FUNCTION_BLOCK "CPG_RecipeSetpoint_STRING"   // FB31617, SCL
TITLE = CPG_RecipeSetpoint_STRING
{ S7_Optimized_Access := 'TRUE' }
AUTHOR : tech.team.motioncontrol@siemens.com
FAMILY : CPG
VERSION : 1.1
// Support: tech.team.motioncontrol@siemens.com
   VAR_INPUT
      enable : Bool;   // If true, setpoint changes are permitted
      disableRecipeControl : Bool;   // If true, the setpoint is no longer handled as a recipe
   END_VAR
   VAR_OUTPUT
      out : String[60];   // Currently running recipe value
      changeEnabled : Bool;   // Enable input is true, setpoint can be changed
      recipeControlDisabled : Bool;   // The value is not subject to recipe controls
      changeNotAllowed : Bool;   // Change is not permitted due to machine state
      recipeSetpointDifference : Bool;   // The currently running (out) value and setpoint value are not equal
   END_VAR
   VAR_IN_OUT
      recipeControl : "CPG_typeRecipeControl";   // Recipe control tag
      recipeSetpoint : "CPG_typeRecipeSetpoint_STRING";   // Recipe setpoint tag
   END_VAR
   VAR
      statFirstScan : Bool := true;
      statPrevChangeNum : Int;
      statPrevSaveNum : Int;
      statPrevCopyNum : Int;
      statPrevDeleteNum : Int;
      statPrevOut : String[60];
      statChangeNotAllowedTimer : TON_TIME;
      statTimerEN : Bool;
   END_VAR
   VAR CONSTANT
      DELAY_TIME : Time := T#3s;
   END_VAR
BEGIN
   //============================================================================================================
   // SIEMENS AG
   // (c)Copyright 2019 All Rights Reserved
   //------------------------------------------------------------------------------------------------------------
   // Library: LCPG
   // Tested with: S7-1500 with FW version V2.1
   // Engineering: TIA Portal V14
   // Restrictions: ---
   // Requirements: S7-1500
   // Functionality: instantiate this once in the program for each recipe setpoint of STRING
   // Support: tech.team.motioncontrol@siemens.com
   //------------------------------------------------------------------------------------------------------------
   // Change log table:
   // Version       Date               Expert in charge    Changes applied
   //  01.01.00     02.01.2019         KB                  Initial Release
   //============================================================================================================
   // Function : CPG_RecipeSetpoint_STRING
   //============================================================================================================

   // Language Selection
   #recipeSetpoint.CurrentSetpointName := #recipeSetpoint.SetpointName[#recipeControl.LanguageSelection];

   //Recipe Disable Control
   #recipeSetpoint.DisableRecipeControl := #disableRecipeControl;

   //Pass through enable bit
   #recipeSetpoint.SetpointChangeEnabled := #enable;

   //Set out value to match initial one on first scan
   IF #statFirstScan THEN
       #recipeSetpoint.CurrentRecipeValue := #recipeSetpoint.RecipeValues[#recipeControl.CurrentRecipeID];
       #recipeSetpoint.OUT := #recipeSetpoint.RecipeValues[#recipeControl.CurrentRecipeID];
       #statFirstScan := false;
   END_IF;


   REGION RECIPE CONTROL
       // Recipe Control - Change, Save, Copy, Delete, Revert setpoint, Save setpoint
       IF NOT (#recipeSetpoint.DisableRecipeControl) THEN
           //Recipe Change command
           IF #recipeControl.RecipeChangeNum <> #statPrevChangeNum THEN
               #recipeSetpoint.OUT := #recipeSetpoint.RecipeValues[#recipeControl.CurrentRecipeID];
               #statPrevChangeNum := #recipeControl.RecipeChangeNum;
               // Prevents multiple commands from being executed if this instruction is not being scanned
               #statPrevSaveNum := #recipeControl.RecipeSaveNum;
               #statPrevCopyNum := #recipeControl.RecipeCopyNum;
               #statPrevDeleteNum := #recipeControl.RecipeDeleteNum;
           END_IF;
           //Recipe Save command
           IF #recipeControl.RecipeSaveNum <> #statPrevSaveNum THEN
               #recipeSetpoint.RecipeValues[#recipeControl.RecipeDestinationID] := #recipeSetpoint.OUT;
               #statPrevSaveNum := #recipeControl.RecipeSaveNum;
               // Prevents multiple commands from being executed if this instruction is not being scanned
               #statPrevCopyNum := #recipeControl.RecipeCopyNum;
               #statPrevDeleteNum := #recipeControl.RecipeDeleteNum;
           END_IF;
           //Recipe Copy command
           IF #recipeControl.RecipeCopyNum <> #statPrevCopyNum THEN
               #recipeSetpoint.RecipeValues[#recipeControl.RecipeDestinationID] := #recipeSetpoint.RecipeValues[#recipeControl.RecipeSourceID];
               #statPrevCopyNum := #recipeControl.RecipeCopyNum;
               // Prevents multiple commands from being executed if this instruction is not being scanned
               #statPrevDeleteNum := #recipeControl.RecipeDeleteNum;
           END_IF;
           //Recipe Delete command
           IF #recipeControl.RecipeDeleteNum <> #statPrevDeleteNum THEN
               //edit this line to change the value a deleted recipe defaults to
               #recipeSetpoint.RecipeValues[#recipeControl.RecipeDestinationID] := ''; 
               #statPrevDeleteNum := #recipeControl.RecipeDeleteNum;
           END_IF;
           //Revert setpoint to saved value
           IF #recipeSetpoint.RevertSetpoint THEN
               #recipeSetpoint.OUT := #recipeSetpoint.RecipeValues[#recipeControl.CurrentRecipeID];
           END_IF;
           //Detect recipe/setpoint difference
           IF (#recipeSetpoint.RecipeValues[#recipeControl.CurrentRecipeID] <> #recipeSetpoint.OUT) AND NOT (#recipeControl.RecipeChange) THEN
               #recipeControl.RecipeSetpointDiff := true;  //signal to recipe control that a setpoint differs
               #recipeSetpoint.RecipeSetpointDiff := true;
           ELSE
               #recipeSetpoint.RecipeSetpointDiff := false;
           END_IF;
           //Save setpoint
           IF #recipeSetpoint.SaveSetpoint THEN
               #recipeSetpoint.RecipeValues[#recipeControl.CurrentRecipeID] := #recipeSetpoint.OUT;
           END_IF;

           //update values stored for current recipe & recipes A, B, & C
           #recipeSetpoint.CurrentRecipeValue := #recipeSetpoint.RecipeValues[#recipeControl.CurrentRecipeID];
           #recipeSetpoint.RecipeValueA := #recipeSetpoint.RecipeValues[#recipeControl.RecipeID_A];
           #recipeSetpoint.RecipeValueB := #recipeSetpoint.RecipeValues[#recipeControl.RecipeID_B];
           #recipeSetpoint.RecipeValueC := #recipeSetpoint.RecipeValues[#recipeControl.RecipeID_C];

       ELSE    //if recipe control is disabled, just update counters
           #recipeSetpoint.RecipeSetpointDiff := false;
           #statPrevChangeNum := #recipeControl.RecipeChangeNum;
           #statPrevSaveNum := #recipeControl.RecipeSaveNum;
           #statPrevCopyNum := #recipeControl.RecipeCopyNum;
           #statPrevDeleteNum := #recipeControl.RecipeDeleteNum;
       END_IF;
   END_REGION


   REGION UPDATE IN VALUE
       //If ENABLE, then changes to the setpoint value are possible
       //otherwise, updating the setpoint is not possible via changing RecipeSetpoint.IN
       IF #enable THEN
           //Clear status bit
           #recipeSetpoint.SetpointChangeDisabled := false;

           // Check for input changed (due to user updating RecipeSetpoint.IN)
           IF (#recipeSetpoint.IN <> #recipeSetpoint.OUT) AND (#recipeSetpoint.OUT = #statPrevOut) THEN
               #recipeSetpoint.OUT := #recipeSetpoint.IN;
           // Check for output changed (due to a recipe change)
           ELSIF (#recipeSetpoint.IN <> #recipeSetpoint.OUT) AND (#recipeSetpoint.OUT <> #statPrevOut) THEN
               #recipeSetpoint.IN := #recipeSetpoint.OUT;
           END_IF;

       ELSE

           // If IN changes, revert and display message
           IF (#recipeSetpoint.IN <> #recipeSetpoint.OUT) OR #recipeSetpoint.RevertSetpoint THEN
               #recipeSetpoint.IN := #recipeSetpoint.OUT;
               #statTimerEN := false;
               #recipeSetpoint.SetpointChangeDisabled := true;
           END_IF;

           //display "setpoint changes not allowed" 3 seconds after inputting an invalid change
           #statChangeNotAllowedTimer(IN := #statTimerEN,
                                  PT := #DELAY_TIME);

           // Continue to display the status bits for the duration of the timer.
           IF #recipeSetpoint.SetpointChangeDisabled THEN
               #statTimerEN := true;
               #recipeSetpoint.SetpointChangeDisabled :=
                   #recipeSetpoint.SetpointChangeDisabled AND #statTimerEN AND NOT #statChangeNotAllowedTimer.Q;
           END_IF;

       END_IF;
   END_REGION


   REGION Set Outputs
       IF (#recipeSetpoint.OUT <> #statPrevOut) THEN
           #statPrevOut := #recipeSetpoint.OUT;
       END_IF;
       #out := #recipeSetpoint.OUT;
       #changeNotAllowed := #recipeSetpoint.SetpointChangeDisabled;
       #recipeSetpointDifference := #recipeSetpoint.RecipeSetpointDiff;
       #recipeControlDisabled := #recipeSetpoint.DisableRecipeControl;
       #changeEnabled := #recipeSetpoint.SetpointChangeEnabled;
   END_REGION

   //  -------------- END OF LOGIC -------------------------
   ENO := TRUE;   // Set the ENO output
END_FUNCTION_BLOCK

FUNCTION "CPG_ModuleInitialize" : Void   // FC31600, SCL
TITLE = CPG_ModuleInitialize
{ S7_Optimized_Access := 'TRUE' }
AUTHOR : tech.team.motioncontrol@siemens.com
FAMILY : CPG
VERSION : 1.0
// Support: tech.team.motioncontrol@siemens.com
   VAR_INPUT
      enableIn : Bool;   // Enable the FB call.
      firstScanBit : Bool;   // Bit used to tell logic that this is the first scan of PLC
   END_VAR
   VAR_IN_OUT
      PackML_ModuleStatus : "CPG_typePackML_ModuleSts";   // PackML Module Status UDT
   END_VAR
BEGIN
   //============================================================================================================
   // SIEMENS AG
   // (c)Copyright 2018 All Rights Reserved
   //------------------------------------------------------------------------------------------------------------
   // Project: CPG Template
   // Tested with: S7-1500 with FW version V2.1
   // Engineering: TIA Portal V14
   // Restrictions: ---
   // Requirements: S7-1500
   // Functionality: This FC will initialize the "PackML" "Status" AND commands within a control module to ensure that the bits are in the correct state IF they are NOT being
   //                used later by that same control module. FOR example, if a start command is NOT being used by a control module, that bit should be turned off TO prevent
   //                unintentional starting OF the machine (in CASE it was accidentally OR through a rung edit turned on). IF a state complete bit FOR a particular state is
   //                NOT being used, that bit should be turned on TO allow the machine TO leave that state. This instruction is NOT needed FOR equipment modules OR the unit
   //                machine since all PackML status AND command bits are programmed in the summation routines.
   // Support: tech.team.motioncontrol@siemens.com
   //------------------------------------------------------------------------------------------------------------
   // Change log table:
   // Version       Date               Expert in charge    Changes applied
   //  01.00.00     01.01.2018         MP                  Initial Release & PackML V1.4  Renamed CPG V1.0
   //  01.01.00     22.05.2018         JP                  Adopted to styleguide
   //============================================================================================================
   // Function : CPG_ModuleInitialize
   //============================================================================================================


   (*  Command vs State Complete:
   •   State complete bits are AND’d together, meaning that all control modules and equipment modules must be done with an acting state 
         before it can transition to the wait state. For example, all of the CM’s and EM’s must be done Stopping before the machine can 
         transition to the Stopped state.
   •   With two exceptions, PackML commands (such as Start, Stop, Abort, Suspend, etc.) are OR’d together, meaning that any 1 control or 
         equipment module can cause the machine to initiate action.  For example, the Stop command initiated from 1 equipment module will 
         stop the entire machine.  

   The only exceptions to this rule are the PackML commands UnHold and UnSuspend.  In either case, the UnHold and UnSuspend commands act 
         like state complete bits.  By doing this in a modular machine architecture, this prevents 1 equipment module from sending the 
         machine into UnHolding or UnSuspending when another equipment module is still wanting the machine to stay held or suspended.  
         For example, assume that both the Infeed Equipment Module (Starved) and Discharge Equipment Module (Blocked) is telling the 
         machine to suspend, if the Infeed Equipment Module has product again, the machine should not UnSuspend without the Discharge 
         Equipment Module also becoming unblocked.
   *)

   IF #firstScanBit OR #enableIn THEN
   // Reset all Command (CMD) bits - this forces the command(CMD) bit to be set in user program if the command is required/used by the CM
       #PackML_ModuleStatus.cmd_Reset           := FALSE; //
       #PackML_ModuleStatus.cmd_Start           := FALSE; //
       #PackML_ModuleStatus.cmd_Stop            := FALSE; //
       #PackML_ModuleStatus.cmd_Hold            := FALSE; //
       #PackML_ModuleStatus.cmd_Suspend         := FALSE; //
       #PackML_ModuleStatus.cmd_Abort           := FALSE; //
       #PackML_ModuleStatus.cmd_Clear           := FALSE; //

   // Set all State Complete (SC) bits - setting the SC bit true allows CM to transition to the next step with no user code need. If the
   // respective SC bit is used by the CM, then user logic must be added to set/reset SC bits as required by the application.
       #PackML_ModuleStatus.sts_Resetting_SC    := TRUE; //
       #PackML_ModuleStatus.sts_Starting_SC     := TRUE; //
       #PackML_ModuleStatus.sts_Stopping_SC     := TRUE; //
       #PackML_ModuleStatus.sts_Holding_SC      := TRUE; //
       #PackML_ModuleStatus.sts_UnHolding_SC    := TRUE; //
       #PackML_ModuleStatus.sts_Suspending_SC   := TRUE; //
       #PackML_ModuleStatus.sts_UnSuspending_SC := TRUE; //
       #PackML_ModuleStatus.sts_Aborting_SC     := TRUE; //
       #PackML_ModuleStatus.sts_Clearing_SC     := TRUE; //
       #PackML_ModuleStatus.sts_Execute_SC      := TRUE; //
       #PackML_ModuleStatus.sts_Completing_SC   := TRUE; //

       //
       #PackML_ModuleStatus.cmd_UnHold          := TRUE; //
       #PackML_ModuleStatus.cmd_UnSuspend       := TRUE; //

   END_IF;  // End "IF FirstScanBit OR EnableIn THEN"

   //  -------------- END OF LOGIC -------------------------
   ENO := TRUE;   // Set the ENO output
END_FUNCTION

FUNCTION "CPG_ArrayLength" : Void   // FC31601, SCL
TITLE = CPG_ArrayLength
{ S7_Optimized_Access := 'TRUE' }
AUTHOR : tech.team.motioncontrol@siemens.com
FAMILY : CPG
VERSION : 1.0
// Support: tech.team.motioncontrol@siemens.com
   VAR_INPUT
      arrayToBeSized : Variant;   // Array to be sized
   END_VAR
   VAR_OUTPUT
      arraySize : Int;   // Number of elements (size) in an array
   END_VAR
BEGIN
   //============================================================================================================
   // SIEMENS AG
   // (c)Copyright 2018 All Rights Reserved
   //------------------------------------------------------------------------------------------------------------
   // Project: CPG Template
   // Tested with: S7-1500 with FW version V2.1
   // Engineering: TIA Portal V14
   // Restrictions: ---
   // Requirements: S7-1x00
   // Functionality: Function Call to determine the length of any array
   //                using optimized S7-1x00 Data Blocks (DB).
   //                This FC can be called from any other FC/FB using any programming
   //                language (SCL, LAD).  Additionally it works with Firmware >= V1.8 
   //                and can determine the size of arrays with elementary (INT,Bool, etc.)
   //                or complex data types (structures)
   // Support: tech.team.motioncontrol@siemens.com
   //------------------------------------------------------------------------------------------------------------
   // Change log table:
   // Version       Date               Expert in charge    Changes applied
   //  01.00.00     08.12.2014         MP                  Initial Release 
   //  01.01.00     22.05.2018         JP                  Adopted to styleguide
   //============================================================================================================
   // Function : CPG_ArrayLength
   //============================================================================================================


   IF IS_ARRAY(#arrayToBeSized) THEN // Check if input is valid array
     #arraySize := UDINT_TO_INT(CountOfElements(#arrayToBeSized)); // Determine the length of the array
   END_IF;

   ENO := TRUE;   // Set the ENO output
END_FUNCTION

// folder: SupportingBlocks/Function_Blocks

FUNCTION_BLOCK "Conveyor"   // FB1, SCL
{ S7_Optimized_Access := 'TRUE' }
VERSION : 0.1
   VAR_INPUT
      bx_PalletSensor : Bool;
      bx_NextReq : Bool;
      bx_PrevReq : Bool;
      ix_CurrentState : DInt;
   END_VAR
   VAR_OUTPUT
      by_ConvFrd : Bool;
      by_NextAck : Bool;
      by_PrevAck : Bool;
      ModuleSts : "CPG_typePackML_ModuleSts";
      iy_SeqStep : Int;
   END_VAR
   VAR
      i_SeqStep : Int;
   END_VAR
BEGIN
   CASE #ix_CurrentState OF
       1://Clearing
           #ModuleSts.sts_Clearing_SC := True;
       2://Stopped
           #ModuleSts.sts_Stopping_SC := False;
           #ModuleSts.sts_Clearing_SC := False;
       3://Starting
           #ModuleSts.sts_Starting_SC := True;
           #iy_SeqStep := #i_SeqStep;
       4://Idle
           #ModuleSts.sts_Resetting_SC := False;
           #by_ConvFrd := False;
           #i_SeqStep := 0;
       5://Suspended
           ;
       6://Execute
           #ModuleSts.sts_Starting_SC := False;
           CASE #i_SeqStep OF
               0://Check if pallet is present
                   IF #bx_PalletSensor AND NOT #bx_PrevReq THEN
                       #i_SeqStep := 2;
                   ELSIF NOT #bx_PalletSensor AND NOT #bx_PrevReq THEN
                       #i_SeqStep := 1;
                   ELSIF #bx_PrevReq THEN
                       #i_SeqStep := 4;
                   END_IF;
               1://Run the conveyor
                   #by_ConvFrd := True;
                   IF #bx_PalletSensor THEN
                       #by_ConvFrd := False;
                       #i_SeqStep := 2;
                   END_IF;
               2://Wait req from next module
                   IF #bx_NextReq THEN
                       #by_NextAck := True;
                       #by_ConvFrd := True;
                       #i_SeqStep := 3;
                   END_IF;
               3://Wait pallet leave
                   IF NOT #bx_PalletSensor THEN
                       #by_NextAck := False;
                       #by_ConvFrd := False;
                       #i_SeqStep := 0;
                   END_IF;
               4://Send the ack to the prev module
                   #by_ConvFrd := True;
                   #by_PrevAck := True;
                   IF #bx_PalletSensor THEN
                       #by_ConvFrd := False;
                       #by_PrevAck := False;
                       #i_SeqStep := 3;
                   END_IF;
           END_CASE;
           //#ModuleSts.sts_Execute_SC := True;
       7://Stopping
           #ModuleSts.sts_Stopping_SC := True;
       8://Aborting
           #ModuleSts.sts_Aborting_SC := True;
       9://Aborted
           #ModuleSts.sts_Aborting_SC := False;
       10://Holding
           #ModuleSts.sts_Holding_SC := True;
       11://Held
           ;
       12://Unholding
           ;
       13://Suspending
           ;
       14://Unsuspending
           ;
       15://Resetting
           #ModuleSts.cmd_Reset := False;
           #ModuleSts.sts_Resetting_SC := True;
       16://Completing
           #ModuleSts.sts_Execute_SC := False;
           #ModuleSts.sts_Completing_SC := True;
       17://Complete
           #ModuleSts.sts_Completing_SC := False;
   END_CASE;
   #iy_SeqStep := #i_SeqStep;
END_FUNCTION_BLOCK

FUNCTION_BLOCK "PackML_Template"   // FB3, SCL
{ S7_Optimized_Access := 'TRUE' }
VERSION : 0.1
   VAR_INPUT
      ix_CurrentState : DInt;
   END_VAR
   VAR_OUTPUT
      ModuleSts : "CPG_typePackML_ModuleSts";
      iy_SeqStep : Int;
   END_VAR
   VAR
      i_SeqStep : Int;
   END_VAR
BEGIN
   CASE #ix_CurrentState OF
       1://Clearing
           #ModuleSts.sts_Clearing_SC := True;
       2://Stopped
           #ModuleSts.sts_Stopping_SC := False;
           #ModuleSts.sts_Clearing_SC := False;
       3://Starting
           #ModuleSts.sts_Starting_SC := True;
           #iy_SeqStep := #i_SeqStep;
       4://Idle
           #ModuleSts.sts_Resetting_SC := False;
           #i_SeqStep := 0;
       5://Suspended
           ;
       6://Execute
           #ModuleSts.sts_Starting_SC := False;
           //#ModuleSts.sts_Execute_SC := True;
       7://Stopping
           #ModuleSts.sts_Stopping_SC := True;
       8://Aborting
           #ModuleSts.sts_Aborting_SC := True;
       9://Aborted
           #ModuleSts.sts_Aborting_SC := False;
       10://Holding
           #ModuleSts.sts_Holding_SC := True;
       11://Held
           ;
       12://Unholding
           ;
       13://Suspending
           ;
       14://Unsuspending
           ;
       15://Resetting
           #ModuleSts.cmd_Reset := False;
           #ModuleSts.sts_Resetting_SC := True;
       16://Completing
           #ModuleSts.sts_Execute_SC := False;
           #ModuleSts.sts_Completing_SC := True;
       17://Complete
           #ModuleSts.sts_Completing_SC := False;
   END_CASE;
   #iy_SeqStep := #i_SeqStep;
END_FUNCTION_BLOCK

FUNCTION_BLOCK "ConveyorCrossing"   // FB4, SCL
{ S7_Optimized_Access := 'TRUE' }
VERSION : 0.1
   VAR_INPUT
      bx_PalletSensor : Bool;
      bx_P1_EmptyPalletReq : Bool;
      bx_P1_ReleasePalletReq : Bool;
      bx_PrevAck : Bool;
      bx_NextAck : Bool;
      ix_CurrentState : DInt;
   END_VAR
   VAR_OUTPUT
      by_RollsFrd : Bool;
      by_RollsRev : Bool;
      by_ChainFrd : Bool;
      by_ChainRev : Bool;
      by_P1_EmptyPalletAck : Bool;
      by_P1_ReleasePalletAck : Bool;
      by_PrevReq : Bool;
      by_NextReq : Bool;
      ModuleSts : "CPG_typePackML_ModuleSts";
      iy_SeqStep : Int;
   END_VAR
   VAR
      i_SeqStep : Int;
   END_VAR
BEGIN
   CASE #ix_CurrentState OF
       1://Clearing
           #ModuleSts.sts_Clearing_SC := True;
       2://Stopped
           #ModuleSts.sts_Stopping_SC := False;
           #ModuleSts.sts_Clearing_SC := False;
       3://Starting
           #ModuleSts.sts_Starting_SC := True;
           #iy_SeqStep := #i_SeqStep;
       4://Idle
           #ModuleSts.sts_Resetting_SC := False;
           #by_ChainFrd := False;
           #by_ChainRev := False;
           #by_RollsFrd := FALSE;
           #by_RollsRev := False;
           #i_SeqStep := 0;
       5://Suspended
           ;
       6://Execute
           #ModuleSts.sts_Starting_SC := False;
           CASE #i_SeqStep OF
               0://Wait req
                   IF #bx_P1_EmptyPalletReq THEN
                       #i_SeqStep := 1;
                   ELSIF #bx_P1_ReleasePalletReq THEN
                       #i_SeqStep := 4;
                   END_IF;
               1://Send the req to the prev module
                   #by_PrevReq := True;
                   IF #bx_PrevAck THEN
                       #i_SeqStep := 2;
                   END_IF;
               2://Start the rolls, wait the empty pallet arrive
                   #by_RollsFrd := True;
                   #by_RollsRev := False;
                   IF #bx_PalletSensor THEN
                       #by_RollsFrd := False;
                       #by_RollsRev := False;
                       #by_PrevReq := False;
                       #i_SeqStep := 3;
                   END_IF;
               3://Start the chain conveyor, wait pallet leave
                   #by_P1_EmptyPalletAck := True;
                   #by_ChainRev := True;
                   #by_ChainFrd := False;
                   IF NOT #bx_PalletSensor AND NOT #bx_P1_EmptyPalletReq THEN
                       #by_ChainRev := False;
                       #by_ChainFrd := False;
                       #i_SeqStep := 0;
                   END_IF;
               4://Send ack to the palletizer, wait pallet arrive at the crossing
                   #by_P1_ReleasePalletAck := True;
                   #by_ChainFrd := True;
                   #by_ChainRev := False;
                   IF #bx_PalletSensor THEN
                       #by_ChainFrd := False;
                       #by_ChainRev := False;
                       #i_SeqStep := 5;
                   END_IF;
               5://Send the req to the next module
                   #by_NextReq := True;
                   IF #bx_NextAck THEN
                       #by_NextReq := False;
                       #i_SeqStep := 6;
                   END_IF;
               6://Start the rolls forward, wait the pallet leave
                   #by_RollsFrd := True;
                   #by_RollsRev := False;
                   IF NOT #bx_PalletSensor THEN
                       #by_RollsFrd := False;
                       #by_RollsRev := False;
                       #i_SeqStep := 0;
                   END_IF;
           END_CASE;
           //#ModuleSts.sts_Execute_SC := True;
       7://Stopping
           #ModuleSts.sts_Stopping_SC := True;
       8://Aborting
           #ModuleSts.sts_Aborting_SC := True;
       9://Aborted
           #ModuleSts.sts_Aborting_SC := False;
       10://Holding
           #ModuleSts.sts_Holding_SC := True;
       11://Held
           ;
       12://Unholding
           ;
       13://Suspending
           ;
       14://Unsuspending
           ;
       15://Resetting
           #ModuleSts.cmd_Reset := False;
           #ModuleSts.sts_Resetting_SC := True;
       16://Completing
           #ModuleSts.sts_Execute_SC := False;
           #ModuleSts.sts_Completing_SC := True;
       17://Complete
           #ModuleSts.sts_Completing_SC := False;
   END_CASE;
   #iy_SeqStep := #i_SeqStep;
END_FUNCTION_BLOCK

FUNCTION_BLOCK "Palletizer"   // FB5, SCL
{ S7_Optimized_Access := 'TRUE' }
VERSION : 0.1
   VAR_INPUT
      bx_BoxSensor : Bool;
      bx_PalletSensor1 : Bool;
      bx_PalletSensor2 : Bool;
      bx_PusherInPos : Bool;
      bx_TrapdoorInPos : Bool;
      bx_PositionerExtended : Bool;
      bx_LiftMoving : Bool;
      bx_BoxReady : Bool;
      bx_PalletReady : Bool;
      bx_ReleasePalletAck : Bool;
      NUMBER_OF_LAYERS : Int;
      ix_CurrentState : DInt;
   END_VAR
   VAR_OUTPUT
      by_BeltFrd : Bool;
      by_BeltRev : Bool;
      by_Pusher : Bool;
      by_Positioner : Bool;
      by_Trapdoor : Bool;
      by_MoveLiftToLimit : Bool;
      by_LiftUp : Bool;
      by_LiftDown : Bool;
      by_ChainFrd : Bool;
      by_ChainRev : Bool;
      by_BoxCam : Bool;
      by_BoxReq : Bool;
      by_PalletReq : Bool;
      by_ReleasePalletReq : Bool;
      ModuleSts : "CPG_typePackML_ModuleSts";
      iy_SeqStep : Int;
      iy_RowCounter : Int;
   END_VAR
   VAR
      i_SeqStep : Int;
      i_RowCounter : Int;
      i_ColumnsCounter : Int;
      i_LayersCounter : Int;
      b_OddLayer : Bool;
      instBoxSensorFTrig : F_TRIG;
      instFullRowOfBoxesTimeout : TON_TIME;
      instLiftTimeout : TON_TIME;
      instPusherTimeout : TON_TIME;
      instTrapdoorTimeout : TON_TIME;
      instLiftDownTimeout : TON_TIME;
   END_VAR
BEGIN
   //----------------------------------------------------------------------------------------
   // Change log table:
   // Version       Date               Expert in charge    Changes applied
   // 1.00          12.03.2022         SGorski             Initial instance of the module
   // 1.01          14.03.2022         SGorski             New timers added
   // 1.02          15.03.2022         SGorski             Now there is a trapdoor reseting in idle step
   //                                                      Odd/Even boxes configurations added
   //                                                      New output added - by_BoxCam
   //                                                      Timers renamed.
   //----------------------------------------------------------------------------------------

   //Falling trigger sensor detection 
   //#instBoxSensorFTrig(CLK := #bx_BoxSensor);


   //Full row of boxes detection timeout
   #instFullRowOfBoxesTimeout(IN := (NOT #b_OddLayer AND #i_RowCounter >= 2) OR (#b_OddLayer AND #i_RowCounter >= 3) ,
                              PT := T#1500ms);

   #instLiftTimeout(IN:=(#i_SeqStep = 4 AND #by_LiftUp)
                      OR (#i_SeqStep = 14 AND #by_LiftDown),
                      PT:=T#500ms);

   #instPusherTimeout(IN := (#i_SeqStep = 7 AND #by_Pusher)
                      OR (#i_SeqStep = 8 AND NOT #by_Pusher),
                      PT := T#1000ms);

   #instTrapdoorTimeout(IN := (#i_SeqStep = 11 AND #by_Trapdoor)
                            OR (#i_SeqStep = 13 AND NOT #by_Trapdoor),
                            PT := T#500ms);

   #instLiftDownTimeout(IN := #i_SeqStep = 12 AND #by_LiftDown,
                        PT := T#1s);



   //Row box counter
   IF #instBoxSensorFTrig.Q OR #bx_BoxSensor THEN
       #i_RowCounter := #i_RowCounter + 1;
   END_IF;



   CASE #ix_CurrentState OF
       1://Clearing
           #ModuleSts.sts_Clearing_SC := True;
       2://Stopped
           #ModuleSts.sts_Stopping_SC := False;
           #ModuleSts.sts_Clearing_SC := False;
       3://Starting
           #ModuleSts.sts_Starting_SC := True;
           #iy_SeqStep := #i_SeqStep;
       4://Idle
           #ModuleSts.sts_Resetting_SC := False;
           #i_SeqStep := 0;
           #by_BeltFrd := false;
           #by_BeltRev := False;
           #by_ChainFrd := False;
           #by_ChainRev := False;
           #by_LiftDown := False;
           #by_LiftUp := False;
           #by_Trapdoor := False;
           #by_MoveLiftToLimit := False;
           #by_Pusher := False;
           #by_Positioner := False;
           #by_BoxReq := False;
           #by_PalletReq := False;
           #by_ReleasePalletReq := False;
           #i_RowCounter := 0;
           #i_ColumnsCounter := 0;
           #i_LayersCounter := 0;
           #b_OddLayer := False;
       5://Suspended
           ;
       6://Execute
           #ModuleSts.sts_Starting_SC := False;
           CASE #i_SeqStep OF
               0://Check if there is a pallet on the chain conveyor   
                   IF #bx_PalletSensor2 THEN
                       #i_SeqStep := 4;
                   ELSE
                       #i_SeqStep := 1;
                   END_IF;
               1://Set the lift fully down
                   #by_MoveLiftToLimit := True;
                   #by_LiftDown := True;
                   #by_LiftUp := False;
                   IF NOT #bx_LiftMoving AND #by_LiftDown AND NOT #by_LiftUp THEN
                       #by_MoveLiftToLimit := False;
                       #by_LiftDown := False;
                       #by_LiftUp := False;
                       #i_SeqStep := 2;
                   END_IF;
               2://Request a new pallet
                   #by_PalletReq := True;
                   IF #bx_PalletReady THEN
                       #i_SeqStep := 3;
                   END_IF;
               3://Start the chain conveyor, wait the pallet arrive
                   #by_ChainFrd := False;
                   #by_ChainRev := True;
                   IF #bx_PalletSensor2 THEN
                       #by_PalletReq := False;
                       #by_ChainFrd := False;
                       #by_ChainRev := False;
                       #i_SeqStep := 4;
                   END_IF;
               4://Set the lift fully up
                   #by_MoveLiftToLimit := True;
                   #by_LiftDown := False;
                   #by_LiftUp := True;
                   IF NOT #bx_LiftMoving AND NOT #by_LiftDown AND #by_LiftUp AND #instLiftTimeout.Q THEN
                       #by_MoveLiftToLimit := False;
                       #by_LiftDown := False;
                       #by_LiftUp := False;
                       #i_SeqStep := 5;
                   END_IF;
               5://Request a new set of boxes
                   #by_BoxReq := True;
                   IF #bx_BoxReady THEN
                       #by_BeltFrd := True;
                       #by_BeltRev := False;
                       #i_SeqStep := 6;
                   END_IF;
               6://Wait the all of the boxes arrive
                   IF #instFullRowOfBoxesTimeout.Q THEN
                       #by_BoxReq := False;
                       #i_SeqStep := 7;
                   END_IF;
               7://Push the boxes onto the trapdoor
                   #by_BeltFrd := False;
                   #by_BeltRev := False;
                   #by_Pusher := True;
                   IF #bx_PusherInPos AND #by_Pusher AND #instPusherTimeout.Q THEN
                       #i_SeqStep := 8;
                   END_IF;
               8://Rectact the pusher and reset the counter
                   #by_Pusher := False;
                   IF #bx_PusherInPos AND NOT #by_Pusher AND #instPusherTimeout.Q THEN
                       #i_RowCounter := 0;
                       #i_ColumnsCounter := #i_ColumnsCounter + 1;
                       IF (NOT #b_OddLayer AND #i_ColumnsCounter >= 3) OR (#b_OddLayer AND #i_ColumnsCounter >= 2) THEN
                           #i_SeqStep := 9;
                       ELSE
                           #i_SeqStep := 5;
                       END_IF;
                   END_IF;
               9://Position the boxes on the trapdoor
                   #by_Positioner := True;
                   IF #bx_PositionerExtended THEN
                       #i_SeqStep := 10;
                   END_IF;
               10://Retract the positioner

                   //IF NOT #bx_PositionerExtended THEN
                       #i_SeqStep := 11;
                  // END_IF;
               11://Open the trapdoor
                   #by_Trapdoor := True;
                   IF #bx_TrapdoorInPos AND #by_Trapdoor AND #instTrapdoorTimeout.Q THEN
                       #i_SeqStep := 12;
                   END_IF;
               12://Move the lift down one layer
                   #by_MoveLiftToLimit := False;
                   #by_LiftDown := True;
                   #by_LiftUp := False;
                   #by_Positioner := False;
                   IF NOT #bx_LiftMoving AND #by_LiftDown AND NOT #by_LiftUp AND #instLiftDownTimeout.Q THEN
                       #i_SeqStep := 13;
                   END_IF;
               13://Close the trapdoor
                   #by_LiftDown := False;
                   #by_LiftUp := False;
                   #by_Trapdoor := False;
                   IF #bx_TrapdoorInPos AND NOT #by_Trapdoor AND #instTrapdoorTimeout.Q THEN
                       #i_ColumnsCounter := 0;
                       #i_LayersCounter := #i_LayersCounter + 1;
                       IF NOT #b_OddLayer THEN
                           #b_OddLayer := True;
                       ELSE
                           #b_OddLayer := False;
                       END_IF;
                       IF #i_LayersCounter >= #NUMBER_OF_LAYERS THEN
                           #i_SeqStep := 14;
                       ELSE
                           #i_SeqStep := 5;
                       END_IF;
                   END_IF;
               14://Move the lift fully down 
                   #by_MoveLiftToLimit := True;
                   #by_LiftDown := True;
                   #by_LiftUp := False;
                   IF NOT #bx_LiftMoving AND #by_LiftDown AND NOT #by_LiftUp AND #instLiftTimeout.Q THEN
                       #by_MoveLiftToLimit := False;
                       #by_LiftDown := False;
                       #by_LiftUp := False;
                       #i_SeqStep := 15;
                   END_IF;
               15://Request the release of the pallet 
                   #by_ReleasePalletReq := True;
                   IF #bx_ReleasePalletAck THEN
                       #i_SeqStep := 16;
                   END_IF;
               16://Move the chain forward
                   #by_ChainFrd := True;
                   #by_ChainRev := False;
                   IF NOT #bx_PalletSensor1 AND NOT #bx_PalletSensor2 THEN
                       #by_ChainFrd := FALSE;
                       #by_ChainRev := False;
                       #by_ReleasePalletReq := False;
                       #i_LayersCounter := 0;
                       #i_SeqStep := 0;
                   END_IF;
           END_CASE;
           //#ModuleSts.sts_Execute_SC := True;
       7://Stopping
           #ModuleSts.sts_Stopping_SC := True;
       8://Aborting
           #ModuleSts.sts_Aborting_SC := True;
       9://Aborted
           #ModuleSts.sts_Aborting_SC := False;
       10://Holding
           #ModuleSts.sts_Holding_SC := True;
       11://Held
           ;
       12://Unholding
           ;
       13://Suspending
           ;
       14://Unsuspending
           ;
       15://Resetting
           #ModuleSts.cmd_Reset := False;
           #ModuleSts.sts_Resetting_SC := True;
       16://Completing
           #ModuleSts.sts_Execute_SC := False;
           #ModuleSts.sts_Completing_SC := True;
       17://Complete
           #ModuleSts.sts_Completing_SC := False;
   END_CASE;
   #iy_SeqStep := #i_SeqStep;
   #iy_RowCounter := #i_RowCounter;
   #by_BoxCam := #b_OddLayer;
END_FUNCTION_BLOCK

FUNCTION_BLOCK "BeltConveyor"   // FB6, SCL
{ S7_Optimized_Access := 'TRUE' }
VERSION : 0.1
   VAR_INPUT
      bx_BoxSensor : Bool;
      bx_BoxReq : Bool;
      ix_CurrentState : DInt;
   END_VAR
   VAR_OUTPUT
      by_BeltFrd : Bool;
      by_BoxReady : Bool;
      ModuleSts : "CPG_typePackML_ModuleSts";
      iy_SeqStep : Int;
   END_VAR
   VAR
      i_SeqStep : Int;
   END_VAR
BEGIN
   CASE #ix_CurrentState OF
       1://Clearing
           #ModuleSts.sts_Clearing_SC := True;
       2://Stopped
           #ModuleSts.sts_Stopping_SC := False;
           #ModuleSts.sts_Clearing_SC := False;
       3://Starting
           #ModuleSts.sts_Starting_SC := True;
           #iy_SeqStep := #i_SeqStep;
       4://Idle
           #ModuleSts.sts_Resetting_SC := False;
           #i_SeqStep := 0;
           #by_BeltFrd := False;
       5://Suspended
           ;
       6://Execute
           #ModuleSts.sts_Starting_SC := False;
           CASE #i_SeqStep OF
               0://Start the conveyor, wait the box arrive
                   #by_BeltFrd := True;
                   IF #bx_BoxSensor THEN
                       #by_BeltFrd := False;
                       #by_BoxReady := True;
                       #i_SeqStep := 1;
                   END_IF;
               1://Wait for the request
                   IF #bx_BoxReq THEN
                       #by_BeltFrd := True;
                       #i_SeqStep := 2;
                   END_IF;
               2://Wait the box leave 
                   IF NOT #bx_BoxSensor THEN
                       #by_BoxReady := False;
                       #i_SeqStep := 0;
                   END_IF;
                   ;
           END_CASE;
           //#ModuleSts.sts_Execute_SC := True;
       7://Stopping
           #ModuleSts.sts_Stopping_SC := True;
       8://Aborting
           #ModuleSts.sts_Aborting_SC := True;
       9://Aborted
           #ModuleSts.sts_Aborting_SC := False;
       10://Holding
           #ModuleSts.sts_Holding_SC := True;
       11://Held
           ;
       12://Unholding
           ;
       13://Suspending
           ;
       14://Unsuspending
           ;
       15://Resetting
           #ModuleSts.cmd_Reset := False;
           #ModuleSts.sts_Resetting_SC := True;
       16://Completing
           #ModuleSts.sts_Execute_SC := False;
           #ModuleSts.sts_Completing_SC := True;
       17://Complete
           #ModuleSts.sts_Completing_SC := False;
   END_CASE;
   #iy_SeqStep := #i_SeqStep;
END_FUNCTION_BLOCK

FUNCTION_BLOCK "FTriggerTest"   // FB7, SCL
{ S7_Optimized_Access := 'TRUE' }
VERSION : 0.1
   VAR_INPUT
      bx_Input : Bool;
      bx_Reset : Bool;
      tx_Timeout : Time;
      ix_CounterMax : Int;
   END_VAR
   VAR_OUTPUT
      by_Output : Bool;
      iy_CounterValue : Int;
   END_VAR
   VAR
      instFTrig : F_TRIG;
      i_Counter : Int;
      instTimeout : TON_TIME;
   END_VAR
BEGIN
   #instFTrig(CLK := #bx_Input);
   #instTimeout(IN := #i_Counter >= #ix_CounterMax,
                PT := T#3s);


   IF #instFTrig.Q THEN
       #i_Counter := #i_Counter + 1;
   END_IF;

   IF #instTimeout.Q THEN
       #by_Output := True;
   END_IF;

   IF #bx_Reset THEN
       #by_Output := False;
   END_IF;


   #iy_CounterValue := #i_Counter;
END_FUNCTION_BLOCK

// folder: SupportingBlocks/LPMLV30_Blocks

FUNCTION_BLOCK "LPMLV30_UnitModeStateManager"   // FB30100, SCL
TITLE = LPMLV30_UnitModeStateManager
{ S7_Optimized_Access := 'TRUE' }
AUTHOR : APC_ERLF
FAMILY : OMAC
// Support: tech.team.motioncontrol@siemens.com 
// Fax: +49 (0) 9131/98-1297
   VAR_INPUT
      UnitMode : DInt := 0;   // Requested unit mode if enableBooleanInterface = FALSE
      UnitModeChangeRequest : Bool := false;   // TRUE: Request unit mode if enableBooleanInterface = FALSE
      CntrlCmd : DInt := 0;   // Request control command if enableBooleanInterface = FALSE
      CmdChangeRequest : Bool := false;   // TRUE: Enable change into requested state if enableBooleanInterface = FALSE
      enableBooleanInterface : Bool := false;   // TRUE: Enable boolean interface
      ProductionModeRequest : Bool := false;   // TRUE: Request change to unit mode Production if enableBooleanInterface = TRUE
      MaintenanceModeRequest : Bool := false;   // TRUE: Request change to unit mode Maintenance if enableBooleanInterface = TRUE
      ManualModeRequest : Bool := false;   // TRUE: Request change to unit mode Manual if enableBooleanInterface = TRUE
      UserMode01Request : Bool := false;   // TRUE: Request change to user-defined unit mode 01 if enableBooleanInterface = TRUE
      UserMode02Request : Bool := false;   // TRUE: Request change to user-defined unit mode 02 if enableBooleanInterface = TRUE
      UserMode03Request : Bool := false;   // TRUE: Request change to user-defined unit mode 03 if enableBooleanInterface = TRUE
      UserMode04Request : Bool := false;   // TRUE: Request change to user-defined unit mode 04 if enableBooleanInterface = TRUE
      UserMode05Request : Bool := false;   // TRUE: Request change to user-defined unit mode 05 if enableBooleanInterface = TRUE
      UserMode06Request : Bool := false;   // TRUE: Request change to user-defined unit mode 06 if enableBooleanInterface = TRUE
      UserMode07Request : Bool := false;   // TRUE: Request change to user-defined unit mode 07 if enableBooleanInterface = TRUE
      UserMode08Request : Bool := false;   // TRUE: Request change to user-defined unit mode 08 if enableBooleanInterface = TRUE
      ResetCmdRequest : Bool := false;   // TRUE: Request control command Reset if enableBooleanInterface = TRUE
      StartCmdRequest : Bool := false;   // TRUE: Request control command Start if enableBooleanInterface = TRUE
      StopCmdRequest : Bool := false;   // TRUE: Request control command Stop if enableBooleanInterface = TRUE
      HoldCmdRequest : Bool := false;   // TRUE: Request control command Hold if enableBooleanInterface = TRUE
      UnholdCmdRequest : Bool := false;   // TRUE: Request control command Unhold if enableBooleanInterface = TRUE
      SuspendCmdRequest : Bool := false;   // TRUE: Request control command Suspend if enableBooleanInterface = TRUE
      UnsuspendCmdRequest : Bool := false;   // TRUE: Request control command Unsuspend if enableBooleanInterface = TRUE
      AbortCmdRequest : Bool := false;   // TRUE: Request control command Abort if enableBooleanInterface = TRUE
      ClearCmdRequest : Bool := false;   // TRUE: Request control command Clear if enableBooleanInterface = TRUE
      CompleteCmdRequest : Bool := false;   // TRUE: Request control command Complete if enableBooleanInterface = TRUE
      SC : Bool := false;   // State change from FALSE to TRUE (rising edge) triggers state complete signal
      configuration : "typeLPMLV30_Configuration";   // FB configuration
   END_VAR
   VAR_OUTPUT
      UnitModeCurrent : DInt := 3;   // Current unit mode
      UnitModeRequested : DInt := 0;   // Requested unit mode
      UnitModeChangeInProcess : Bool := false;   // Unit mode change in process
      StateCurrent : DInt := 2;   // Current state
      StateRequested : DInt := 0;   // Requested state
      StateChangeInProcess : Bool := false;   // State change in process
      ProductionModeActive : Bool := false;   // TRUE: Unit mode Production is currently active
      MaintenanceModeActive : Bool := false;   // TRUE: Unit mode Maintenance is currently active
      ManualModeActive : Bool := false;   // TRUE: Unit mode Manual is currently active
      UserMode01Active : Bool := false;   // TRUE: User-defined unit mode 01 is currently active
      UserMode02Active : Bool := false;   // TRUE: User-defined unit mode 02 is currently active
      UserMode03Active : Bool := false;   // TRUE: User-defined unit mode 03 is currently active
      UserMode04Active : Bool := false;   // TRUE: User-defined unit mode 04 is currently active
      UserMode05Active : Bool := false;   // TRUE: User-defined unit mode 05 is currently active
      UserMode06Active : Bool := false;   // TRUE: User-defined unit mode 06 is currently active
      UserMode07Active : Bool := false;   // TRUE: User-defined unit mode 07 is currently active
      UserMode08Active : Bool := false;   // TRUE: User-defined unit mode 08 is currently active
      ClearingStateActive : Bool := false;   // TRUE: State Clearing is currently active
      StoppedStateActive : Bool := false;   // TRUE: State Stopped is currently active
      StartingStateActive : Bool := false;   // TRUE: State Starting is currently active
      IdleStateActive : Bool := false;   // TRUE: State Idle is currently active
      SuspendedStateActive : Bool := false;   // TRUE: State Suspended is currently active
      ExecuteStateActive : Bool := false;   // TRUE: State Execute is currently active
      StoppingStateActive : Bool := false;   // TRUE: State Stopping is currently active
      AbortingStateActive : Bool := false;   // TRUE: State Aborting is currently active
      AbortedStateActive : Bool := false;   // TRUE: State Aborted is currently active
      HoldingStateActive : Bool := false;   // TRUE: State Holding is currently active
      HeldStateActive : Bool := false;   // TRUE: State Held is currently active
      UnholdingStateActive : Bool := false;   // TRUE: State Unholding is currently active
      SuspendingStateActive : Bool := false;   // TRUE: State Suspending is currently active
      UnsuspendingStateActive : Bool := false;   // TRUE: State Unsuspending is currently active
      ResettingStateActive : Bool := false;   // TRUE: State Resetting is currently active
      CompletingStateActive : Bool := false;   // TRUE: State Completing is currently active
      CompleteStateActive : Bool := false;   // TRUE: State Complete is currently active
      StatesDisabled : DInt;   // Disabled states in current unit mode
      diagnostics : "typeLPMLV30_Diagnostics";   // Diagnostics information of FB
   END_VAR
   VAR
      statConfiguration : "typeLPMLV30_Configuration";   // FB configuration
      statUnitModeChangeRequest : Bool := false;   // TRUE: Enable change into requested unit mode
      statCmdChangeRequest : Bool := false;   // TRUE: Enable change into requested state
      statFirstCycle : Bool := true;   // First cycle of run
      statSCOld : Bool := false;   // For edge detection
      statUnitMode : DInt := 3;   // Current command mode
      statUnitModeOld : DInt := 3;   // For edge detection
      statUnitModeCurrentInternal : DInt := 3;   // Current internal Mode
      statUnitModeCurrentInternalOld : DInt := 0;   // For edge detection
      statStateCurrentOld : DInt := 2;   // For edge detection
      statStateInternal : DInt := 2;   // Current internal state
      statStateInternalOld : DInt := 0;   // For edge detection
      statCntrlCmdOld : DInt := 0;   // For edge detection
      statStatesInCurrentMode : Struct   // Copied from configuration
         clearing : Bool;
         stopped : Bool;
         starting : Bool;
         idle : Bool;
         suspended : Bool;
         execute : Bool;
         stopping : Bool;
         aborting : Bool;
         aborted : Bool;
         holding : Bool;
         held : Bool;
         unholding : Bool;
         suspending : Bool;
         unsuspending : Bool;
         resetting : Bool;
         completing : Bool;
         complete : Bool;
      END_STRUCT;
      statBooleanInterfaceModeOld : DWord;   // For edge detection
      statBooleanInterfaceCmdOld : Word;   // For edge detection
      statCmdChangeRequestOld : Bool := false;   // For edge detection
      statUnitModeChangeRequestOld : Bool := false;   // For edge detection
   END_VAR
   VAR_TEMP
      tempCntrlCmd : DInt;   // Temporary control command
      tempBooleanInterfaceMode : DWord;   // Status of boolean Mode inputs if boolean interface is active